(* Logix 5000 project; controller MV vendor 1 type 14 code 217 rev 31.11; software revision 31.00; part 36 of 53 *)
(* tags used below, declared in another part *)
   Alarm_Reset : BOOL;
   Analog_Fault_No : DINT;
   Analog_Simulation_Enabled : BOOL;
   CWD : CHECKWORD_FLAGS;
   Default_Check_Time : DINT;
   Dummy : BOOL;
   MV_Copy_from_fv_file : INT;
   MV_Copy_to_fv_file : INT;
   MV_MV20_LTX07_AI : PlantItem;   // MV20_LTX07
   MV_MV20_LTX07_AI_RawInput : ALIAS FOR Remote_IO:10:I.Ch03Data;   // Real Analog Input , Do Not Use In Code
   MV_MV20_LTX07_TrueLevel : REAL;
   MV_MV20_LTX07_TruePressure : REAL;
   MV_MV20_PTX01_AI : PlantItem;   // MV20_PTX01
   MV_MV20_PTX01_AI_RawInput : ALIAS FOR Remote_IO:10:I.Ch00Data;   // Real Analog Input , Do Not Use In Code
   MV_MV21_LTX07_AI : PlantItem;   // MV21_LTX07
   MV_MV21_LTX07_AI_RawInput : ALIAS FOR Remote_IO:10:I.Ch04Data;   // Real Analog Input , Do Not Use In Code
   MV_MV21_LTX07_TrueLevel : REAL;
   MV_MV21_LTX07_TruePressure : REAL;
   MV_MV21_PTX01_AI : PlantItem;   // MV21_PTX01
   MV_MV21_PTX01_AI_RawInput : ALIAS FOR Remote_IO:10:I.Ch01Data;   // Real Analog Input , Do Not Use In Code
   MV_MV22_LTX07_AI : PlantItem;   // MV22_LTX07
   MV_MV22_LTX07_AI_RawInput : ALIAS FOR Remote_IO:10:I.Ch05Data;   // Real Analog Input , Do Not Use In Code
   MV_MV22_LTX07_TrueLevel : REAL;
   MV_MV22_LTX07_TruePressure : REAL;
   MV_MV22_PTX01_AI : PlantItem;   // MV22_PTX01
   MV_MV22_PTX01_AI_RawInput : ALIAS FOR Remote_IO:10:I.Ch02Data;   // Real Analog Input , Do Not Use In Code
   MV_N106 : INT[255];   // ROUSE_BUFF Rouser control vesse l data buffer
   MV_N110 : INT[255];   // MV DATA 0 CURRENT FV DATA
   MV_N111 : INT[50];   // MV 1, CURRENT FV DATA
   MV_N112 : INT[50];   // MV 2, CURRENT FV DATA
   MV_N113 : INT[50];   // MV 3, CURRENT FV DATA
   MV_N114 : INT[50];   // MV 4, CURRENT FV DATA
   MV_N115 : INT[50];   // MV 5, CURRENT FV DATA
   MV_N116 : INT[50];   // MV 6, CURRENT FV DATA
   MV_N117 : INT[50];   // MV 7, CURRENT FV DATA
   MV_N118 : INT[50];   // MV 8, CURRENT FV DATA
   MV_N119 : INT[50];   // MV 9, CURRENT FV DATA
   MV_N120 : INT[50];   // MV 10, CURRENT FV DATA
   MV_N121 : INT[50];   // MV 11, CURRENT FV DATA
   MV_N122 : INT[50];   // MV 12, CURRENT FV DATA
   MV_N123 : INT[50];   // MV 13, CURRENT FV DATA
   MV_N124 : INT[50];   // MV 14, CURRENT FV DATA
   MV_N125 : INT[50];   // MV 15, CURRENT FV DATA
   MV_N126 : INT[50];   // MV 16, CURRENT FV DATA
   MV_N127 : INT[50];   // MV 17, CURRENT FV DATA
   MV_N128 : INT[50];   // MV 18, CURRENT FV DATA
   MV_N129 : INT[50];   // MV 19, CURRENT FV DATA
   MV_N130 : INT[50];   // MV 30, CURRENT FV DATA
   MV_N131 : INT[50];   // MV 31, CURRENT FV DATA
   One_Second_One_Scan : ALIAS FOR One_Second_1_scan;
   overrange_RIO_analog_value : REAL;
   underrange_RIO_analog_value : REAL;
(* MV_Common, continued *)

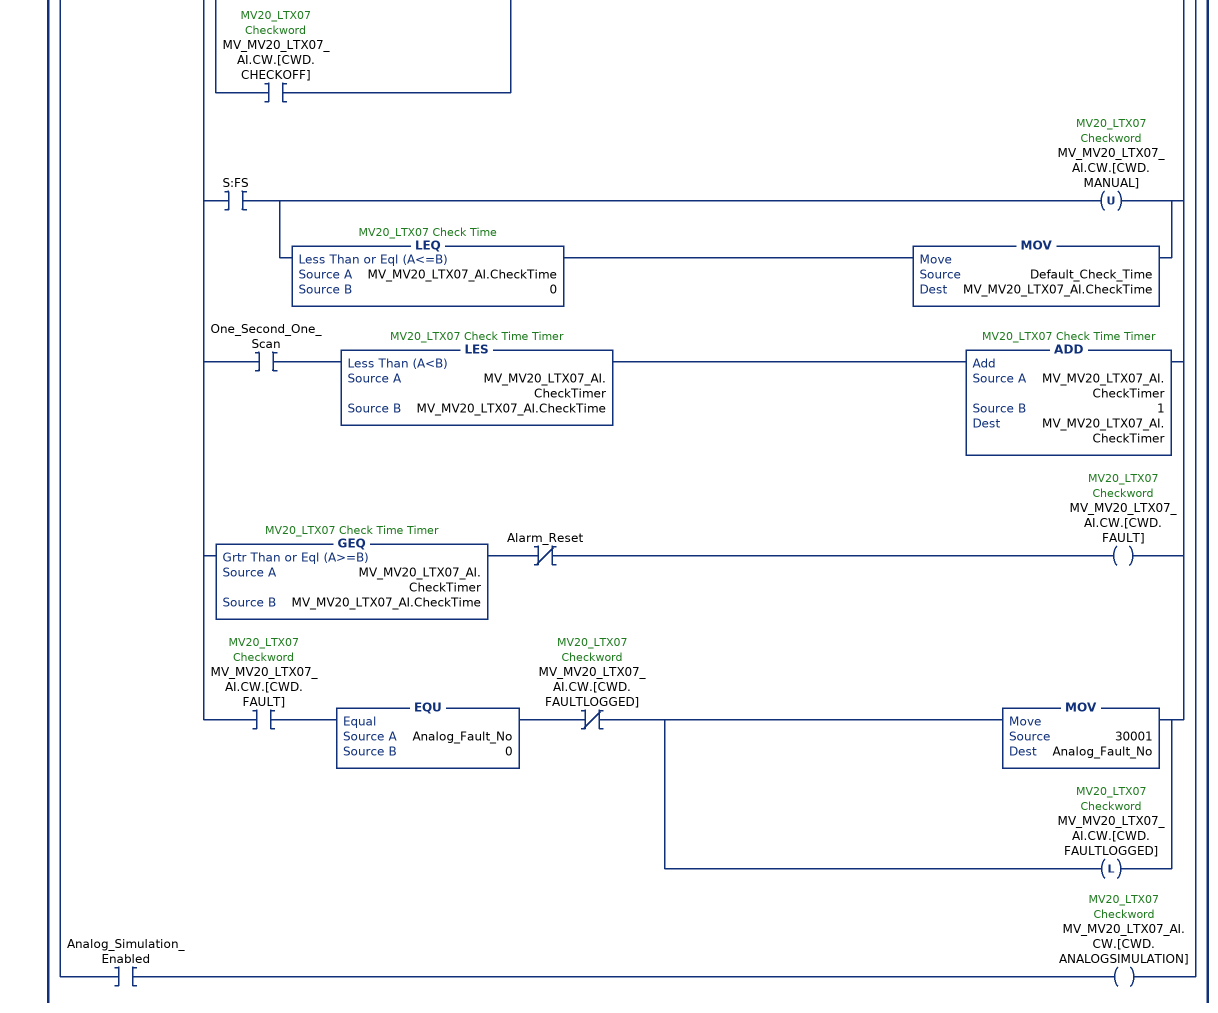
   [picture p835: MV_Common/MV_Analogs rungs 41-41]
   41: [XIO(Analog_Simulation_Enabled) [XIO(MV_MV20_LTX07_AI.CW.[CWD.MANUAL]) [JSR(Analog_Scale_ItoF,5,MV_MV20_LTX07_AI_RawInput,4000.0,20000.0,0.0,29.0,MV_MV20_LTX07_AI.Scaled) ,GRT(MV_MV20_PTX01_AI.Scaled,0) GRT(MV_MV20_LTX07_AI.Scaled,MV_MV20_PTX01_AI.Scaled) SUB(MV_MV20_LTX07_AI.Scaled,MV_MV20_PTX01_AI.Scaled,MV_MV20_LTX07_TruePressure) ,LEQ(MV_MV20_PTX01_AI.Scaled,0) GRT(MV_MV20_LTX07_AI.Scaled,MV_MV20_PTX01_AI.Scaled) MOV(MV_MV20_LTX07_AI.Scaled,MV_MV20_LTX07_TruePressure) ,LEQ(MV_MV20_LTX07_AI.Scaled,MV_MV20_PTX01_AI.Scaled) MOV(0,MV_MV20_LTX07_TruePressure) ,JSR(Analog_scale_ftof,5,MV_MV20_LTX07_TruePressure,0.0,5.743,0.0,260.0,MV_MV20_LTX07_TrueLevel) ,LEQ(MV_MV20_LTX07_TrueLevel,0) MOV(0,MV_MV20_LTX07_TrueLevel) ] ,MOV(MV_MV20_LTX07_AI_RawInput,MV_MV20_LTX07_AI.RawInput) ,[LIM(underrange_RIO_analog_value,MV_MV20_LTX07_AI_RawInput,overrange_RIO_analog_value) ,XIC(MV_MV20_LTX07_AI.CW.[CWD.CHECKOFF]) ] CLR(MV_MV20_LTX07_AI.CheckTimer) ,XIC(S:FS) [OTU(MV_MV20_LTX07_AI.CW.[CWD.MANUAL]) ,LEQ(MV_MV20_LTX07_AI.CheckTime,0) MOV(Default_Check_Time,MV_MV20_LTX07_AI.CheckTime) ] ,XIC(One_Second_One_Scan) LES(MV_MV20_LTX07_AI.CheckTimer,MV_MV20_LTX07_AI.CheckTime) ADD(MV_MV20_LTX07_AI.CheckTimer,1,MV_MV20_LTX07_AI.CheckTimer) ,GEQ(MV_MV20_LTX07_AI.CheckTimer,MV_MV20_LTX07_AI.CheckTime) XIO(Alarm_Reset) OTE(MV_MV20_LTX07_AI.CW.[CWD.FAULT]) ,XIC(MV_MV20_LTX07_AI.CW.[CWD.FAULT]) EQU(Analog_Fault_No,0) XIO(MV_MV20_LTX07_AI.CW.[CWD.FAULTLOGGED]) [MOV(30001,Analog_Fault_No) ,OTL(MV_MV20_LTX07_AI.CW.[CWD.FAULTLOGGED]) ] ] ,XIC(Analog_Simulation_Enabled) OTE(MV_MV20_LTX07_AI.CW.[CWD.ANALOGSIMULATION]) ];
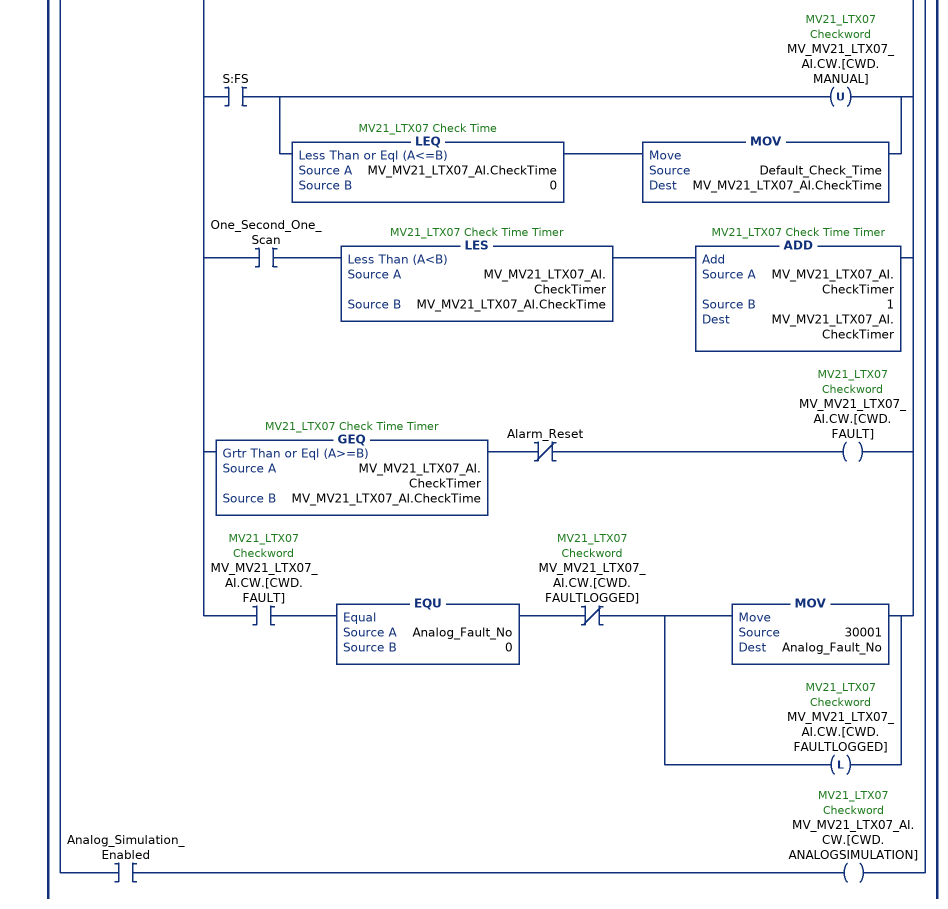
   42: [XIO(Analog_Simulation_Enabled) [XIO(MV_MV21_LTX07_AI.CW.[CWD.MANUAL]) [JSR(Analog_Scale_ItoF,5,MV_MV21_LTX07_AI_RawInput,4000.0,20000.0,0.0,29.0,MV_MV21_LTX07_AI.Scaled) ,GRT(MV_MV21_PTX01_AI.Scaled,0) SUB(MV_MV21_LTX07_AI.Scaled,MV_MV21_PTX01_AI.Scaled,MV_MV21_LTX07_TruePressure) ,LEQ(MV_MV21_PTX01_AI.Scaled,0) MOV(MV_MV21_LTX07_AI.Scaled,MV_MV21_LTX07_TruePressure) ,JSR(Analog_scale_ftof,5,MV_MV21_LTX07_TruePressure,0.0,5.743,0.0,260.0,MV_MV21_LTX07_TrueLevel) ,LEQ(MV_MV21_LTX07_TrueLevel,0) MOV(0,MV_MV21_LTX07_TrueLevel) ] ,MOV(MV_MV21_LTX07_AI_RawInput,MV_MV21_LTX07_AI.RawInput) ,[LIM(underrange_RIO_analog_value,MV_MV21_LTX07_AI_RawInput,overrange_RIO_analog_value) ,XIC(MV_MV21_LTX07_AI.CW.[CWD.CHECKOFF]) ] CLR(MV_MV21_LTX07_AI.CheckTimer) ,XIC(S:FS) [OTU(MV_MV21_LTX07_AI.CW.[CWD.MANUAL]) ,LEQ(MV_MV21_LTX07_AI.CheckTime,0) MOV(Default_Check_Time,MV_MV21_LTX07_AI.CheckTime) ] ,XIC(One_Second_One_Scan) LES(MV_MV21_LTX07_AI.CheckTimer,MV_MV21_LTX07_AI.CheckTime) ADD(MV_MV21_LTX07_AI.CheckTimer,1,MV_MV21_LTX07_AI.CheckTimer) ,GEQ(MV_MV21_LTX07_AI.CheckTimer,MV_MV21_LTX07_AI.CheckTime) XIO(Alarm_Reset) OTE(MV_MV21_LTX07_AI.CW.[CWD.FAULT]) ,XIC(MV_MV21_LTX07_AI.CW.[CWD.FAULT]) EQU(Analog_Fault_No,0) XIO(MV_MV21_LTX07_AI.CW.[CWD.FAULTLOGGED]) [MOV(30001,Analog_Fault_No) ,OTL(MV_MV21_LTX07_AI.CW.[CWD.FAULTLOGGED]) ] ] ,XIC(Analog_Simulation_Enabled) OTE(MV_MV21_LTX07_AI.CW.[CWD.ANALOGSIMULATION]) ];
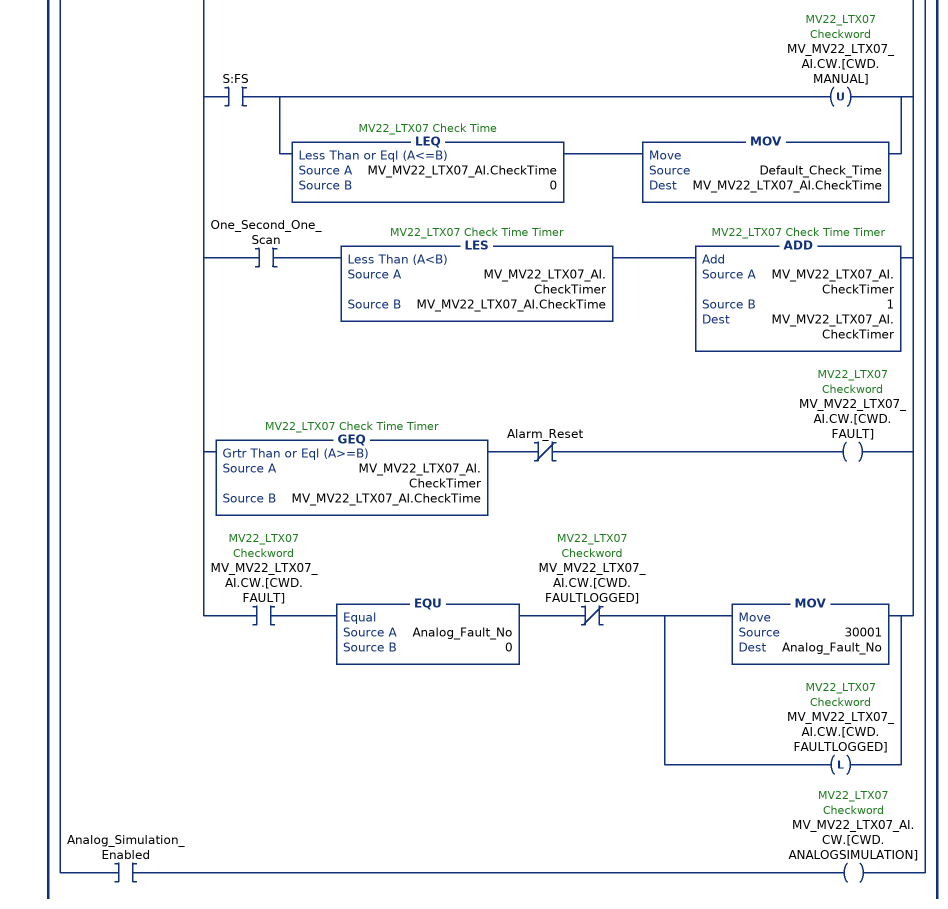
   43: [XIO(Analog_Simulation_Enabled) [XIO(MV_MV22_LTX07_AI.CW.[CWD.MANUAL]) [JSR(Analog_Scale_ItoF,5,MV_MV22_LTX07_AI_RawInput,4000.0,20000.0,0.0,29.0,MV_MV22_LTX07_AI.Scaled) ,GRT(MV_MV22_PTX01_AI.Scaled,0) SUB(MV_MV22_LTX07_AI.Scaled,MV_MV22_PTX01_AI.Scaled,MV_MV22_LTX07_TruePressure) ,LEQ(MV_MV22_PTX01_AI.Scaled,0) MOV(MV_MV22_LTX07_AI.Scaled,MV_MV22_LTX07_TruePressure) ,JSR(Analog_scale_ftof,5,MV_MV22_LTX07_TruePressure,0.0,5.743,0.0,260.0,MV_MV22_LTX07_TrueLevel) ,LEQ(MV_MV22_LTX07_TrueLevel,0) MOV(0,MV_MV22_LTX07_TrueLevel) ] ,MOV(MV_MV22_LTX07_AI_RawInput,MV_MV22_LTX07_AI.RawInput) ,[LIM(underrange_RIO_analog_value,MV_MV22_LTX07_AI_RawInput,overrange_RIO_analog_value) ,XIC(MV_MV22_LTX07_AI.CW.[CWD.CHECKOFF]) ] CLR(MV_MV22_LTX07_AI.CheckTimer) ,XIC(S:FS) [OTU(MV_MV22_LTX07_AI.CW.[CWD.MANUAL]) ,LEQ(MV_MV22_LTX07_AI.CheckTime,0) MOV(Default_Check_Time,MV_MV22_LTX07_AI.CheckTime) ] ,XIC(One_Second_One_Scan) LES(MV_MV22_LTX07_AI.CheckTimer,MV_MV22_LTX07_AI.CheckTime) ADD(MV_MV22_LTX07_AI.CheckTimer,1,MV_MV22_LTX07_AI.CheckTimer) ,GEQ(MV_MV22_LTX07_AI.CheckTimer,MV_MV22_LTX07_AI.CheckTime) XIO(Alarm_Reset) OTE(MV_MV22_LTX07_AI.CW.[CWD.FAULT]) ,XIC(MV_MV22_LTX07_AI.CW.[CWD.FAULT]) EQU(Analog_Fault_No,0) XIO(MV_MV22_LTX07_AI.CW.[CWD.FAULTLOGGED]) [MOV(30001,Analog_Fault_No) ,OTL(MV_MV22_LTX07_AI.CW.[CWD.FAULTLOGGED]) ] ] ,XIC(Analog_Simulation_Enabled) OTE(MV_MV22_LTX07_AI.CW.[CWD.ANALOGSIMULATION]) ];
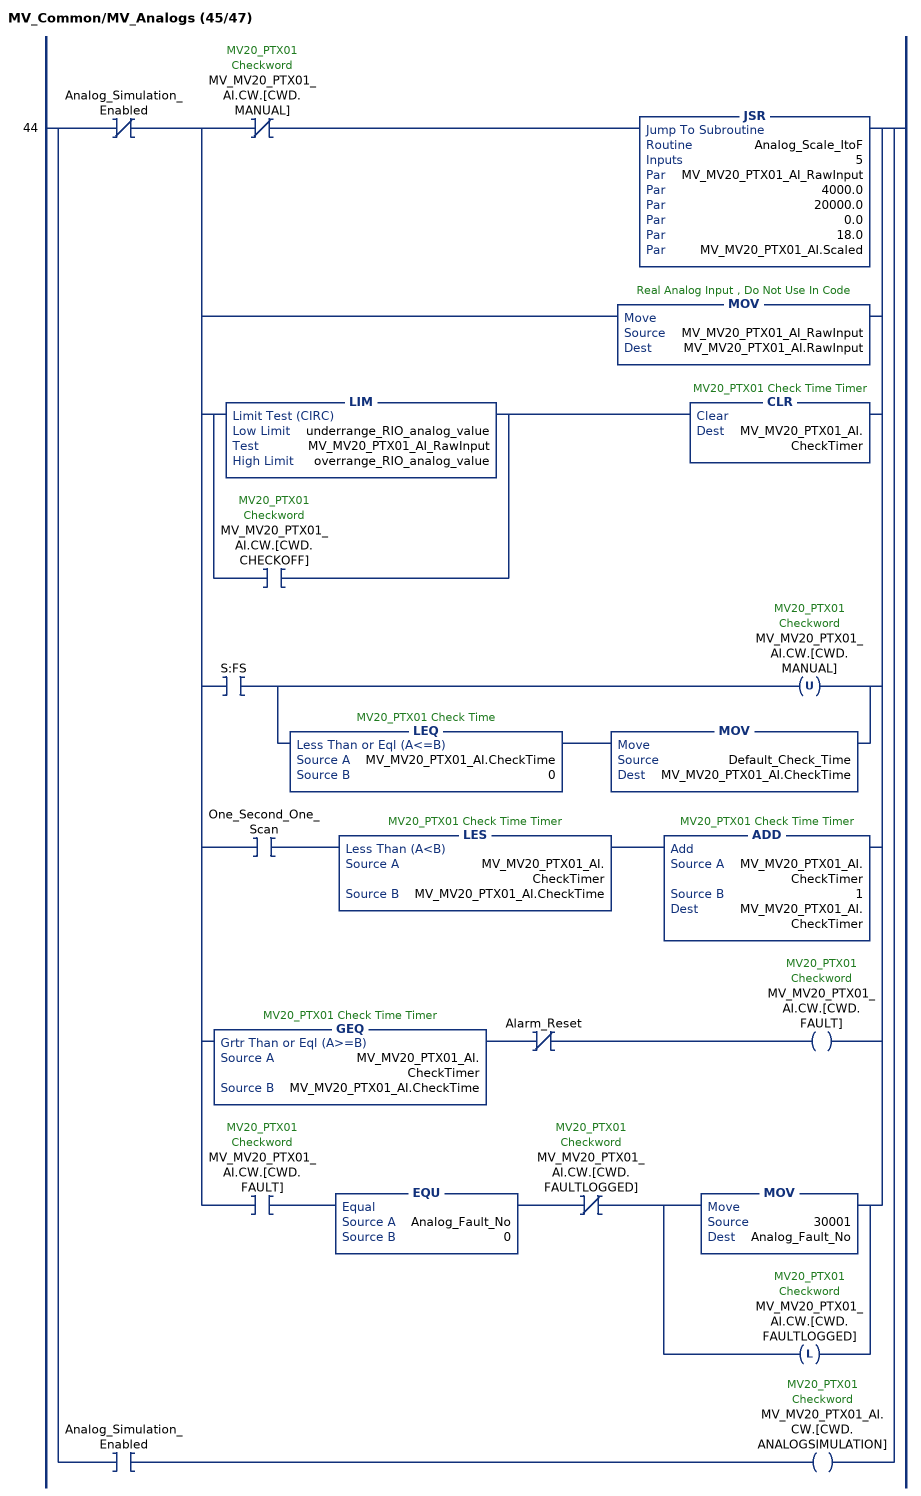
   44: [XIO(Analog_Simulation_Enabled) [XIO(MV_MV20_PTX01_AI.CW.[CWD.MANUAL]) JSR(Analog_Scale_ItoF,5,MV_MV20_PTX01_AI_RawInput,4000.0,20000.0,0.0,18.0,MV_MV20_PTX01_AI.Scaled) ,MOV(MV_MV20_PTX01_AI_RawInput,MV_MV20_PTX01_AI.RawInput) ,[LIM(underrange_RIO_analog_value,MV_MV20_PTX01_AI_RawInput,overrange_RIO_analog_value) ,XIC(MV_MV20_PTX01_AI.CW.[CWD.CHECKOFF]) ] CLR(MV_MV20_PTX01_AI.CheckTimer) ,XIC(S:FS) [OTU(MV_MV20_PTX01_AI.CW.[CWD.MANUAL]) ,LEQ(MV_MV20_PTX01_AI.CheckTime,0) MOV(Default_Check_Time,MV_MV20_PTX01_AI.CheckTime) ] ,XIC(One_Second_One_Scan) LES(MV_MV20_PTX01_AI.CheckTimer,MV_MV20_PTX01_AI.CheckTime) ADD(MV_MV20_PTX01_AI.CheckTimer,1,MV_MV20_PTX01_AI.CheckTimer) ,GEQ(MV_MV20_PTX01_AI.CheckTimer,MV_MV20_PTX01_AI.CheckTime) XIO(Alarm_Reset) OTE(MV_MV20_PTX01_AI.CW.[CWD.FAULT]) ,XIC(MV_MV20_PTX01_AI.CW.[CWD.FAULT]) EQU(Analog_Fault_No,0) XIO(MV_MV20_PTX01_AI.CW.[CWD.FAULTLOGGED]) [MOV(30001,Analog_Fault_No) ,OTL(MV_MV20_PTX01_AI.CW.[CWD.FAULTLOGGED]) ] ] ,XIC(Analog_Simulation_Enabled) OTE(MV_MV20_PTX01_AI.CW.[CWD.ANALOGSIMULATION]) ];
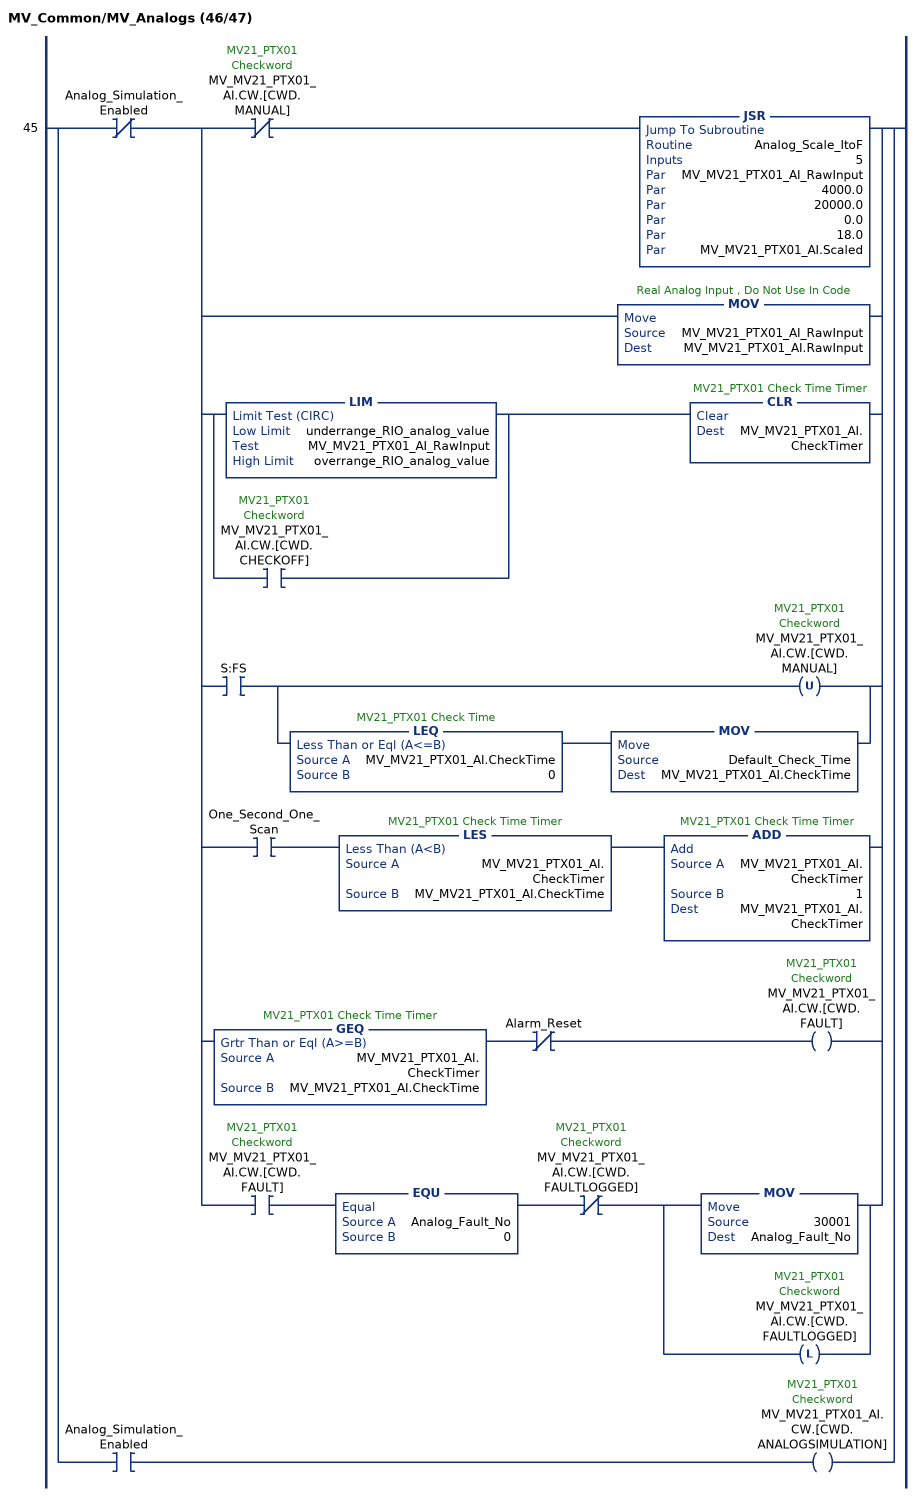
   45: [XIO(Analog_Simulation_Enabled) [XIO(MV_MV21_PTX01_AI.CW.[CWD.MANUAL]) JSR(Analog_Scale_ItoF,5,MV_MV21_PTX01_AI_RawInput,4000.0,20000.0,0.0,18.0,MV_MV21_PTX01_AI.Scaled) ,MOV(MV_MV21_PTX01_AI_RawInput,MV_MV21_PTX01_AI.RawInput) ,[LIM(underrange_RIO_analog_value,MV_MV21_PTX01_AI_RawInput,overrange_RIO_analog_value) ,XIC(MV_MV21_PTX01_AI.CW.[CWD.CHECKOFF]) ] CLR(MV_MV21_PTX01_AI.CheckTimer) ,XIC(S:FS) [OTU(MV_MV21_PTX01_AI.CW.[CWD.MANUAL]) ,LEQ(MV_MV21_PTX01_AI.CheckTime,0) MOV(Default_Check_Time,MV_MV21_PTX01_AI.CheckTime) ] ,XIC(One_Second_One_Scan) LES(MV_MV21_PTX01_AI.CheckTimer,MV_MV21_PTX01_AI.CheckTime) ADD(MV_MV21_PTX01_AI.CheckTimer,1,MV_MV21_PTX01_AI.CheckTimer) ,GEQ(MV_MV21_PTX01_AI.CheckTimer,MV_MV21_PTX01_AI.CheckTime) XIO(Alarm_Reset) OTE(MV_MV21_PTX01_AI.CW.[CWD.FAULT]) ,XIC(MV_MV21_PTX01_AI.CW.[CWD.FAULT]) EQU(Analog_Fault_No,0) XIO(MV_MV21_PTX01_AI.CW.[CWD.FAULTLOGGED]) [MOV(30001,Analog_Fault_No) ,OTL(MV_MV21_PTX01_AI.CW.[CWD.FAULTLOGGED]) ] ] ,XIC(Analog_Simulation_Enabled) OTE(MV_MV21_PTX01_AI.CW.[CWD.ANALOGSIMULATION]) ];
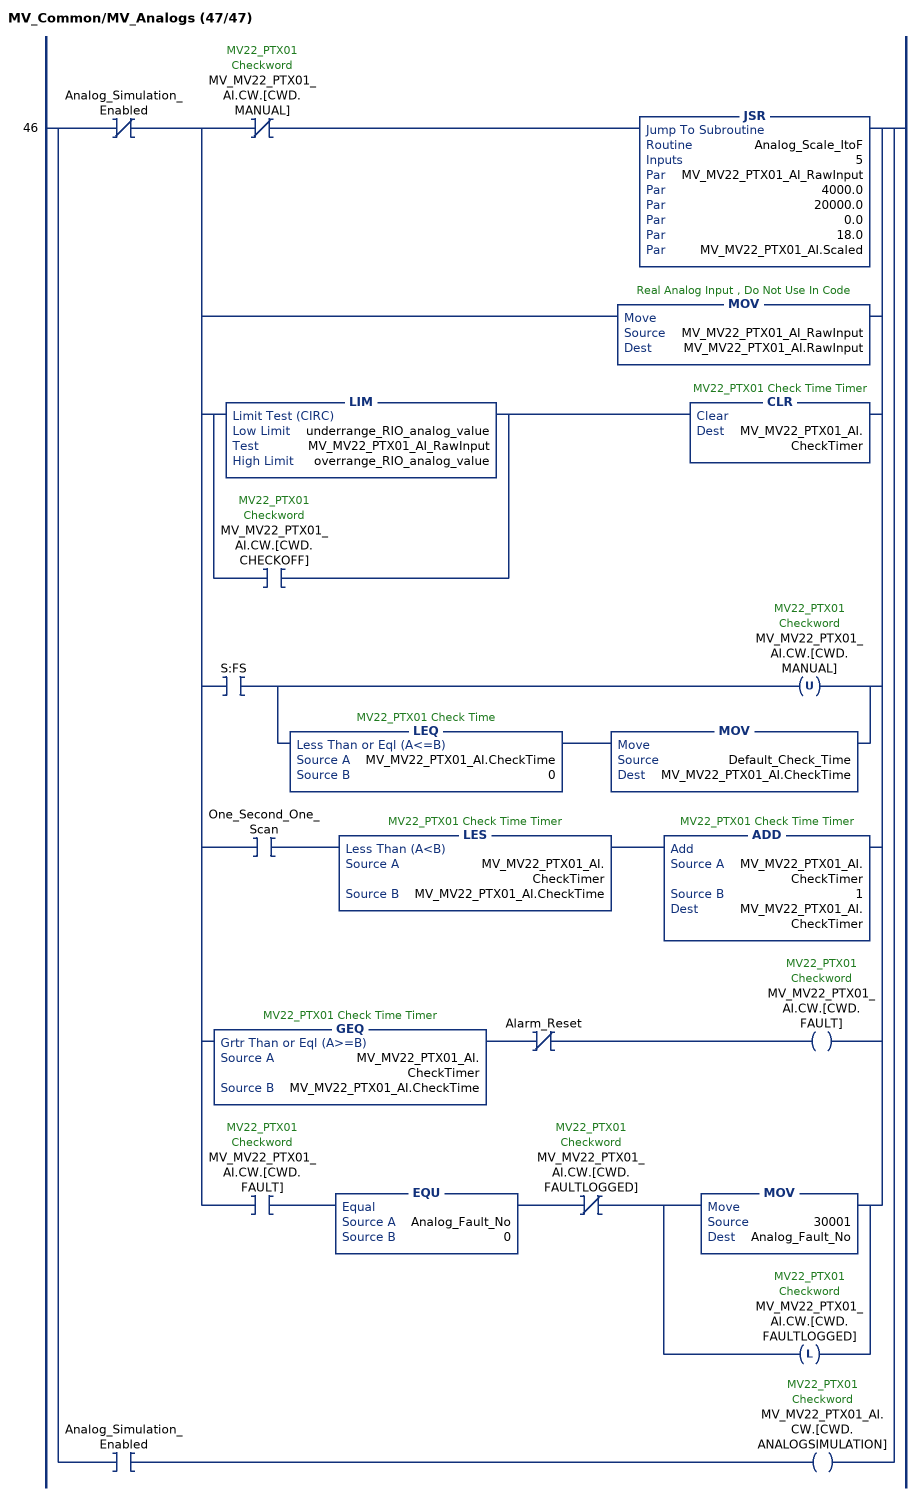
   46: [XIO(Analog_Simulation_Enabled) [XIO(MV_MV22_PTX01_AI.CW.[CWD.MANUAL]) JSR(Analog_Scale_ItoF,5,MV_MV22_PTX01_AI_RawInput,4000.0,20000.0,0.0,18.0,MV_MV22_PTX01_AI.Scaled) ,MOV(MV_MV22_PTX01_AI_RawInput,MV_MV22_PTX01_AI.RawInput) ,[LIM(underrange_RIO_analog_value,MV_MV22_PTX01_AI_RawInput,overrange_RIO_analog_value) ,XIC(MV_MV22_PTX01_AI.CW.[CWD.CHECKOFF]) ] CLR(MV_MV22_PTX01_AI.CheckTimer) ,XIC(S:FS) [OTU(MV_MV22_PTX01_AI.CW.[CWD.MANUAL]) ,LEQ(MV_MV22_PTX01_AI.CheckTime,0) MOV(Default_Check_Time,MV_MV22_PTX01_AI.CheckTime) ] ,XIC(One_Second_One_Scan) LES(MV_MV22_PTX01_AI.CheckTimer,MV_MV22_PTX01_AI.CheckTime) ADD(MV_MV22_PTX01_AI.CheckTimer,1,MV_MV22_PTX01_AI.CheckTimer) ,GEQ(MV_MV22_PTX01_AI.CheckTimer,MV_MV22_PTX01_AI.CheckTime) XIO(Alarm_Reset) OTE(MV_MV22_PTX01_AI.CW.[CWD.FAULT]) ,XIC(MV_MV22_PTX01_AI.CW.[CWD.FAULT]) EQU(Analog_Fault_No,0) XIO(MV_MV22_PTX01_AI.CW.[CWD.FAULTLOGGED]) [MOV(30001,Analog_Fault_No) ,OTL(MV_MV22_PTX01_AI.CW.[CWD.FAULTLOGGED]) ] ] ,XIC(Analog_Simulation_Enabled) OTE(MV_MV22_PTX01_AI.CW.[CWD.ANALOGSIMULATION]) ];
END_ROUTINE

ROUTINE MV_Copy_Vessel_File   (* ladder *)
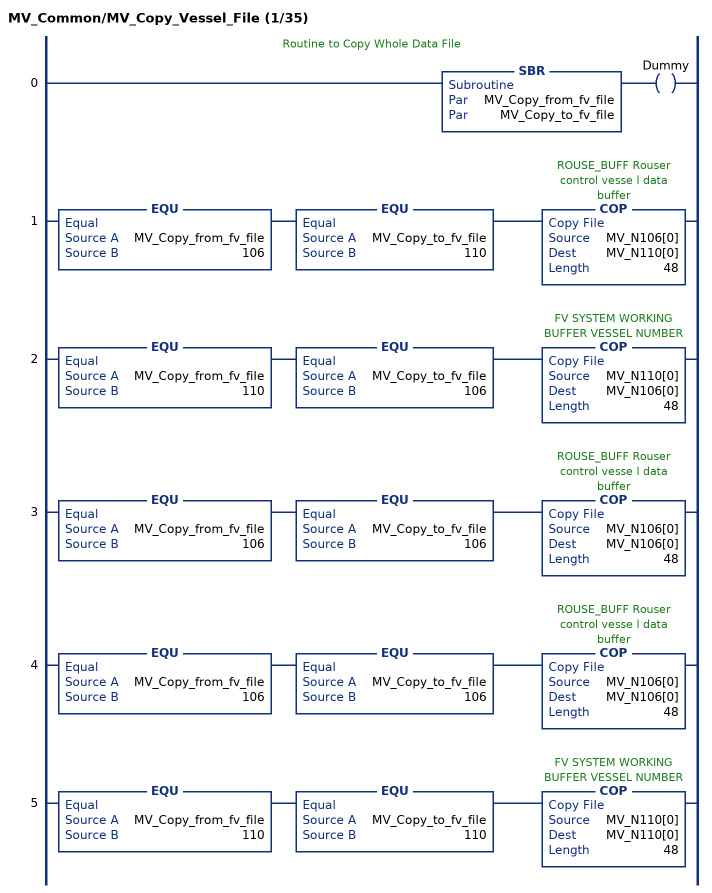
   // Routine to Copy Whole Data File
   0: SBR(MV_Copy_from_fv_file,MV_Copy_to_fv_file)OTE(Dummy);
   1: EQU(MV_Copy_from_fv_file,106)EQU(MV_Copy_to_fv_file,110)COP(MV_N106[0],MV_N110[0],48);
   2: EQU(MV_Copy_from_fv_file,110)EQU(MV_Copy_to_fv_file,106)COP(MV_N110[0],MV_N106[0],48);
   3: EQU(MV_Copy_from_fv_file,106)EQU(MV_Copy_to_fv_file,106)COP(MV_N106[0],MV_N106[0],48);
   4: EQU(MV_Copy_from_fv_file,106)EQU(MV_Copy_to_fv_file,106)COP(MV_N106[0],MV_N106[0],48);
   5: EQU(MV_Copy_from_fv_file,110)EQU(MV_Copy_to_fv_file,110)COP(MV_N110[0],MV_N110[0],48);